
FUNCTION "SCALE_D" : Real   // FC334, SCL
TITLE = SCALE_D
{ S7_Optimized_Access := 'FALSE' }
AUTHOR : hugo
FAMILY : SIGPRO
NAME : SCALED
VERSION : 1.2
// Scale_D is used to translate and scale a DWORD input x to a real output.
// the input is limited to I_LO <= X <= I_HI.
   VAR_INPUT
      X : DWord;
      I_LO : DWord;
      I_HI : DWord;
      O_LO : Real;
      O_HI : Real;
   END_VAR
BEGIN


     IF #I_HI = #I_LO THEN
       #SCALE_D := #O_LO;
     ELSE
       #SCALE_D := (#O_HI - #O_LO) / DINT_TO_REAL(DWORD_TO_DINT(#I_HI) - DWORD_TO_DINT(#I_LO))
                  * DINT_TO_REAL(LIMIT(MN:=DWORD_TO_DINT(#I_LO),IN:=DWORD_TO_DINT(#X),MX:=DWORD_TO_DINT(#I_HI)) 
                  - DWORD_TO_DINT(#I_LO)) + #O_LO;
     END_IF;


   (* revision history
   hm  18. may. 2008 rev 1.0
     original version

   hm  13. nov. 2008 rev 1.1
     corrected formula for negative gradient

   hm  11. jan 2011  rev 1.2
     avoid division by 0
   *)
END_FUNCTION

FUNCTION "SCALE_R" : Real   // FC335, SCL
TITLE = SCALE_R
{ S7_Optimized_Access := 'FALSE' }
AUTHOR : hugo
FAMILY : SIGPRO
NAME : SCALER
VERSION : 1.2
// Scale_R is used to translate and scale a REAL input x to a real output.
// the input is limited to I_LO <= X <= I_HI.
   VAR_INPUT
      X : Real;
      I_LO : Real;
      I_HI : Real;
      O_LO : Real;
      O_HI : Real;
   END_VAR
BEGIN


     IF #I_LO = #I_HI THEN
       #SCALE_R := #O_LO;
     ELSE
       #SCALE_R := (#O_HI - #O_LO) / (#I_HI - #I_LO) * (LIMIT(MN:=#I_LO,IN:=#X,MX:=#I_HI) - #I_LO) + #O_LO;
     END_IF;


   (* revision history
   hm  18. may. 2008 rev 1.0
     original version

   hm  13. nov. 2008 rev 1.1
     corrected formula for negative gradient

   hm  11. jan 2011  rev 1.2
     avoid division by 0

   *)
END_FUNCTION

FUNCTION "SCALE_X2" : Real   // FC336, SCL
TITLE = SCALE_X2
{ S7_Optimized_Access := 'FALSE' }
AUTHOR : hugo
FAMILY : SIGPRO
NAME : SCALEX2
VERSION : 1.1
// this functiob block can scale up to two inputs.
// the input can select between two ues with true or false.
// the summed output is then scaled by an scale input K and a offset O can be added to the output.
// the min and max input configurations can be edited in the cfc editor by double clicking the symbol body.
   VAR_INPUT
      IN1 : Bool;
      IN2 : Bool;
      K : Real;
      O : Real;
      IN1_MIN : Real;
      IN1_MAX : Real;
      IN2_MIN : Real;
      IN2_MAX : Real;
   END_VAR
BEGIN


   #SCALE_X2 := (SEL(G:=#IN1,IN0:=#IN1_MIN, IN1:=#IN1_MAX)+ 
                SEL(G:=#IN2,IN0:=#IN2_MIN, IN1:=#IN2_MAX))*#K + #O;


   (* revision history
   hm  19. jan, 2007   rev 1.0
       original version

   hm  26. oct. 2008   rev 1.1
       code optimized

   *)
END_FUNCTION

FUNCTION "SCALE_X4" : Real   // FC337, SCL
TITLE = SCALE_X4
{ S7_Optimized_Access := 'FALSE' }
AUTHOR : hugo
FAMILY : SIGPRO
NAME : SCALEX4
VERSION : 1.0
// this function can scale up to 4 inputs.
// the input can select between two ues with true or false.
// the summed output is then scaled by an scale input K and a offset O can be added to the output.
// the min and max input configurations can be edited in the cfc editor by double clicking the symbol body.
   VAR_INPUT
      in1 : Bool;
      in2 : Bool;
      in3 : Bool;
      in4 : Bool;
      K : Real;
      O : Real;
      in1_min : Real;
      in1_max : Real;
      in2_min : Real;
      in2_max : Real;
      in3_min : Real;
      in3_max : Real;
      in4_min : Real;
      in4_max : Real;
   END_VAR
BEGIN


     IF NOT #in1 THEN #SCALE_X4 := #in1_min; ELSE #SCALE_X4 := #in1_max; END_IF;
     IF NOT #in2 THEN #SCALE_X4 := #SCALE_X4 + #in2_min; ELSE #SCALE_X4 := #SCALE_X4 + #in2_max; END_IF;
     IF NOT #in3 THEN #SCALE_X4 := #SCALE_X4 + #in3_min; ELSE #SCALE_X4 := #SCALE_X4 + #in3_max; END_IF;
     IF NOT #in4 THEN #SCALE_X4 := #SCALE_X4 + #in4_min; ELSE #SCALE_X4 := #SCALE_X4 + #in4_max; END_IF;
     #SCALE_X4 := #SCALE_X4 * #K + #O;

   (* revision history

   *)
END_FUNCTION

FUNCTION "SCALE_X8" : Real   // FC338, SCL
TITLE = SCALE_X8
{ S7_Optimized_Access := 'FALSE' }
AUTHOR : hugo
FAMILY : SIGPRO
NAME : SCALEX8
VERSION : 1.2
// this function can scale up to 4 inputs.
// the input can select between two ues with true or false.
// the summed output is then scaled by an scale input K and a offset O can be added to the output.
// the min and max input configurations can be edited in the cfc editor by double clicking the symbol body.
   VAR_INPUT
      in1 : Bool;
      in2 : Bool;
      in3 : Bool;
      in4 : Bool;
      in5 : Bool;
      in6 : Bool;
      in7 : Bool;
      in8 : Bool;
      K : Real;
      O : Real;
      in1_min : Real;
      in1_max : Real;
      in2_min : Real;
      in2_max : Real;
      in3_min : Real;
      in3_max : Real;
      in4_min : Real;
      in4_max : Real;
      in5_min : Real;
      in5_max : Real;
      in6_min : Real;
      in6_max : Real;
      in7_min : Real;
      in7_max : Real;
      in8_min : Real;
      in8_max : Real;
   END_VAR
BEGIN


   #SCALE_X8 := (SEL(G:=#in1,IN0:=#in1_min,IN1:=#in1_max) + 
                SEL(G:=#in2,IN0:=#in2_min,IN1:=#in2_max) + 
                SEL(G:=#in3,IN0:=#in3_min,IN1:=#in3_max) + 
                SEL(G:=#in4,IN0:=#in4_min,IN1:=#in4_max) +
                SEL(G:=#in5,IN0:=#in5_min,IN1:=#in5_max) + 
                SEL(G:=#in6,IN0:=#in6_min,IN1:=#in6_max) + 
                SEL(G:=#in7,IN0:=#in7_min,IN1:=#in7_max) + 
                SEL(G:=#in8,IN0:=#in8_min,IN1:=#in8_max))* #K + #O;


   (* revision history
   hm  19. jan. 2008   rev 1.0
       original version

   hm  26. oct. 2008   rev 1.1
       optimized code

   hm  24. jan. 2008   rev 1.2
       corrected error in formula
   *)
END_FUNCTION

FUNCTION "STAIR" : Real   // FC339, SCL
TITLE = STAIR
{ S7_Optimized_Access := 'FALSE' }
AUTHOR : oscat
FAMILY : SIGPRO
NAME : STAIR
VERSION : 1.4
// the function stair converts an anlog input signal to a staircase like output.
// D is the step width for the output signal.
// if D = 0 then the output follows the input without a chage.
   VAR_INPUT
      X : Real;
      D : Real;
   END_VAR
BEGIN


   IF #D > 0.0 THEN
       #STAIR := DINT_TO_REAL(REAL_TO_DINT(#X / #D)) * #D;
   ELSE
       #STAIR := #X;
   END_IF;


   (* revision history
   hm  28 jan 2007     rev 1.0
       original version

   hm  27 dec 2007     rev 1.1
       changed code for better performance

   hm  6. jan 2008     rev 1.2
       further performance improvement

   hm  26. oct. 2008       rev 1.3
       optimized code

   hm  10. mar. 2009   rev 1.4
       real constants updated to new systax using dot

   *)
END_FUNCTION

FUNCTION "WORD_TO_RANGE" : Real   // FC340, SCL
TITLE = WORD_TO_RANGE
{ S7_Optimized_Access := 'FALSE' }
AUTHOR : hugo
FAMILY : SIGPRO
NAME : WO2RA
VERSION : 1.1
// Word_to_Range converts a Byte into a real between low and high.
   VAR_INPUT
      X : Word;
      low : Real;
      high : Real;
   END_VAR
BEGIN


   #WORD_TO_RANGE := (#high - #low) * DINT_TO_REAL(WORD_TO_DINT(#X)) * 0.00001525902189669640 + #low;


   (* revision history
   hm  9. jan 2008 rev 1.0
       original version

   hm  10. mar. 2009   rev 1.1
       improved code
   *)
END_FUNCTION

// ===== PLC "Engineering automation"  Unspecific CPU S7 300 =====

VAR_GLOBAL CONSTANT   // PLC tag table "STEP7 classic symbols"
   "debug" : Bool := FALSE;
   "N" : Int := 0;
   "offset" : Int := 0;
   "one" : Byte := 16#01;
   "offset_1" : DWord := 0;
END_VAR

DATA_BLOCK "IDB_STIME"   // DB64
{ S7_Optimized_Access := 'FALSE' }
AUTHOR : dalbi
FAMILY : MEASURE
VERSION : 0.0
// stored: InstanceOfName STIME
"STIME"
BEGIN
END_DATA_BLOCK

FUNCTION_BLOCK "STIME"   // FB64, SCL
TITLE = STIME
{ S7_Optimized_Access := 'FALSE' }
AUTHOR : dalbi
FAMILY : MEASURE
NAME : STIME
VERSION : 1.4
// this function block makes sure that the timer of a siemens sps counts from 0 - 2^32-1.
   VAR_OUTPUT
      tx : DWord;
      at_tx AT tx : Array[0..31] of Bool;
   END_VAR
   VAR
      last_time : DWord;
      bit31 : Bool;
      init : Bool := TRUE;
   END_VAR
   VAR_TEMP
      TOP_SI : Struct
         EV_CLASS : Byte;
         EV_NUM : Byte;
         PRIORITY : Byte;
         NUM : Byte;
         TYP2_3 : Byte;
         TYP1 : Byte;
         ZI1 : Word;
         ZI2_3 : DWord;
      END_STRUCT;
      START_UP_SI : Struct
         EV_CLASS : Byte;
         EV_NUM : Byte;
         PRIORITY : Byte;
         NUM : Byte;
         TYP2_3 : Byte;
         TYP1 : Byte;
         ZI1 : Word;
         ZI2_3 : DWord;
      END_STRUCT;
      ERR : Int;
   END_VAR
BEGIN


   (* this FB is only necessary for siemens sps
   the siemens sps timer counts from 0 to 2^31-1 and starts at 0 sfter overrun.
   this means that the bit 31 (the highest bit ) will never be used and therefore
   a problem arises when t2 - t1 is checked.
   t2 - t1 is always valid also in an timer overrun situation where the time t1 is very high and t2 is very low.
   the result of the subtraction t2 - t1 however is still valid.
   this calculation does not work for soiemens because the highest bit is not used.

   this module stores the highest bit, changes the highest bit at every overrun occurence and stuffs ther highest bit in the output.
   the output is then used by t_plc_us and t_plc_ms.

   the correction needs and fb and not a function because the value of the highest bit has to be stored.

   do never use this function block in a codesys environment. the timer in codesys is correct and runs from 0 to 2^32-1
   *)

   (* read actual startup info *)
   (* OB1_SCAN_1  BYTE  -  B#16#01: Abschluss des Neustarts (Warmstarts)
                        -  B#16#02: Abschluss des Wiederanlaufs
                        -  B#16#03: Abschluss des freien Zyklus
                        -  B#16#04: Abschluss des Kaltstarts
                        -  B#16#05: Erster OB 1-Zyklus der neuen Master-CPU nach 
                                    Master-Reserve-Umschaltung und STOP des 
                                    bisherigen Masters *)

   #ERR := RD_SINFO (TOP_SI => #TOP_SI, START_UP_SI => #START_UP_SI);

   (* reset last_time on system startup *)
   IF #TOP_SI.EV_NUM = 1 OR #TOP_SI.EV_NUM = 2 OR #TOP_SI.EV_NUM = 4 OR NOT #init THEN 
       #last_time := 0;
       #bit31 := false;
       #init := true;
   END_IF;

   (* read the system timer *)
   #tx := DINT_TO_DWORD(T_CONV(TIME_TCK()));

   (* check for overrun *)
   IF DWORD_TO_DINT(#tx) < DWORD_TO_DINT(#last_time) THEN
       (* an overrun has occured, change the value of the highest bit *)
       #bit31 := NOT #bit31;
   END_IF;

   (* stuff the highest bit into the timer value *)
   #at_tx[7] := #bit31;

   (* remember the last system time for the next overrun check *)
   #last_time := #tx;


   (* revision history
   DA  14.9.2007 rev 1.0
     original version

   DA  24.2.2008 rev 1.1
     added self reset on system startup

   DA   2.5.2008 rev 1.2
     corect a problem running under OB35

   DA  12.3.2009 rev 1.3
     corect a problem run on different CPUs

   DA  22.12.2009 rev 1.4
     corect a problem on startup
   *)
END_FUNCTION_BLOCK

FUNCTION_BLOCK "TP_1D"   // FB68, SCL
TITLE = TP_1D
{ S7_Optimized_Access := 'FALSE' }
AUTHOR : hugo
FAMILY : GENERAT
NAME : TP_1D
VERSION : 1.0
// TP_2 generates a pulse every time it is calles with in := TRUE.
// the module will reset IN by itself so no clearing of in is necessary.
// in addition the timer can be cleared asynchronously with rst.
// also the rst input is cleared by the module itself.
// the timer can be retriggered as often as necessary. it will count PT from the last trigger.
// after the time PT1 is elapsed, the timer blocks itself for PT2 and only allow new sequences after PT2 has elapsed.
// 
// uses: T_PLC_MS [FC64]
//       STIME [FB64],IDB_STIME [DB64]
   VAR_INPUT
      IN : Bool;
      PT1 : Time;
      PTD : Time;
      RST : Bool;
   END_VAR
   VAR_OUTPUT
      Q : Bool;
      W : Bool;
   END_VAR
   VAR
      tx : Time;
      start : Time;
      ix : Bool;
   END_VAR
BEGIN


   (* read system timer *)
   #tx := T_CONV(DWORD_TO_DINT("T_PLC_MS"()));

   IF #RST THEN
       #Q := FALSE;
       #RST := FALSE;
       #W := FALSE;
   ELSIF #W THEN
       IF #tx - #start >= #PTD THEN
           #W := FALSE;
       END_IF;
   ELSIF #IN AND NOT #ix THEN
       #Q := TRUE;
       #start := #tx;
       #IN := FALSE;
   ELSIF #tx - #start >= #PT1 THEN
       #Q := FALSE;
       #W := TRUE;
       #start := #tx;
   END_IF;

   #ix := #IN;



   (* revision history
   hm  28. jun. 2008
       original version

   *)
END_FUNCTION_BLOCK

FUNCTION_BLOCK "TC_S"   // FB134, SCL
TITLE = TC_S
{ S7_Optimized_Access := 'FALSE' }
AUTHOR : hugo
FAMILY : MEASURE
NAME : TC_S
VERSION : 1.2
// TC_S delivers the time it was last called on the output TC in seconds.
// 
// uses: T_PLC_US [FC65]
//       STIME [FB64],IDB_STIME [DB64]
   VAR_OUTPUT
      TC : Real;
   END_VAR
   VAR
      init : Bool;
      tx : DWord;
      last : DWord;
   END_VAR
   VAR_TEMP
      TOP_SI : Struct
         EV_CLASS : Byte;
         EV_NUM : Byte;
         PRIORITY : Byte;
         NUM : Byte;
         TYP2_3 : Byte;
         TYP1 : Byte;
         ZI1 : Word;
         ZI2_3 : DWord;
      END_STRUCT;
      START_UP_SI : Struct
         EV_CLASS : Byte;
         EV_NUM : Byte;
         PRIORITY : Byte;
         NUM : Byte;
         TYP2_3 : Byte;
         TYP1 : Byte;
         ZI1 : Word;
         ZI2_3 : DWord;
      END_STRUCT;
      ERR : Int;
   END_VAR
BEGIN


   (* read actual startup info *)
   (* OB1_SCAN_1  BYTE  -  B#16#01: Abschluss des Neustarts (Warmstarts)
                        -  B#16#02: Abschluss des Wiederanlaufs
                        -  B#16#03: Abschluss des freien Zyklus
                        -  B#16#04: Abschluss des Kaltstarts
                        -  B#16#05: Erster OB 1-Zyklus der neuen Master-CPU nach 
                                    Master-Reserve-Umschaltung und STOP des 
                                    bisherigen Masters *)

     #ERR := RD_SINFO (TOP_SI => #TOP_SI, START_UP_SI => #START_UP_SI);

   (* reset last_time on system startup *)
   IF #TOP_SI.EV_NUM = 1 OR #TOP_SI.EV_NUM = 2 OR #TOP_SI.EV_NUM = 4 THEN 
       #last := 0;
       #init := FALSE;
   END_IF;

   (* read system timer *)
   #tx := "T_PLC_US"();

   IF NOT #init THEN
       #init := TRUE;
       #TC := 0.0;
   ELSE
       #TC := (DINT_TO_REAL(DWORD_TO_DINT(#tx)) - DINT_TO_REAL(DWORD_TO_DINT(#last)))*1.0E-6;
   END_IF;
   #last := #tx;


   (* revision history
   hm  13. mar. 2008   rev 1.0
       original version

   hm  16. mar 2008    rev 1.1
       added type conversion to avoid warnings under codesys 3.0

   hm  11. mar. 2009   rev 1.2
       changed real constants to use dot syntax

   *)
END_FUNCTION_BLOCK

FUNCTION_BLOCK "DRIVER_1"   // FB202, SCL
TITLE = DRIVER_1
{ S7_Optimized_Access := 'FALSE' }
AUTHOR : hugo
FAMILY : AUTOMAT
NAME : DRIVER_1
VERSION : 1.0
// driver_1 is a multi purpose driver.
// a rising edge in in sets the output high if toggle is flase. while toggle is true, a rising edge on in toggles the output Q.
// if a timeout is specified the output q will be reset to false automatically after the timeout has elapsed.
// a asynchronous reset and set will force the output high or low respectively.
   VAR_INPUT
      Toggle_Mode : Bool;
      Timeout : Time;
      SET : Bool;
      IN : Bool;
      RST : Bool;
   END_VAR
   VAR_OUTPUT
      Q : Bool;
   END_VAR
   VAR
      off : TON;
      edge : Bool;
   END_VAR
BEGIN


     IF #off.Q THEN #Q := FALSE; END_IF;
     IF #RST THEN
       #Q := FALSE;
     ELSIF #SET THEN
       #Q := TRUE;
     ELSIF #IN AND NOT #edge THEN
       IF #Toggle_Mode THEN #Q := NOT #Q; ELSE #Q := TRUE; END_IF;
     END_IF;
     #edge := #IN;
     IF #Timeout > t#0s THEN #off(IN := #Q, PT := #Timeout); END_IF;


   (* revision history
   hm  2. jan 2008   rev 1.0
     original version

   *)
END_FUNCTION_BLOCK

FUNCTION_BLOCK "DRIVER_4"   // FB203, SCL
TITLE = DRIVER_4
{ S7_Optimized_Access := 'FALSE' }
AUTHOR : hugo
FAMILY : AUTOMAT
NAME : DRIVER_4
VERSION : 1.0
// driver_1 is a multi purpose driver.
// a rising edge in in sets the output high if toggle is flase. while toggle is true, a rising edge on in toggles the output Q.
// if a timeout is specified the output q will be reset to false automatically after the timeout has elapsed.
// a asynchronous reset and set will force the output high or low respectively.
// 
// uses: DRIVER_1 [FB202]
   VAR_INPUT
      Toggle_Mode : Bool;
      Timeout : Time;
      SET : Bool;
      IN0 : Bool;
      IN1 : Bool;
      IN2 : Bool;
      IN3 : Bool;
      RST : Bool;
   END_VAR
   VAR_OUTPUT
      Q0 : Bool;
      Q1 : Bool;
      Q2 : Bool;
      Q3 : Bool;
   END_VAR
   VAR
      d0 : "DRIVER_1";
      d1 : "DRIVER_1";
      d2 : "DRIVER_1";
      d3 : "DRIVER_1";
   END_VAR
BEGIN


     #d0(SET:=#SET, IN:=#IN0, RST:=#RST, Toggle_Mode:=#Toggle_Mode, Timeout:=#Timeout);
     #d1(SET:=#SET, IN:=#IN1, RST:=#RST, Toggle_Mode:=#Toggle_Mode, Timeout:=#Timeout);
     #d2(SET:=#SET, IN:=#IN2, RST:=#RST, Toggle_Mode:=#Toggle_Mode, Timeout:=#Timeout);
     #d3(SET:=#SET, IN:=#IN3, RST:=#RST, Toggle_Mode:=#Toggle_Mode, Timeout:=#Timeout);
     #Q0 := #d0.Q;
     #Q1 := #d1.Q;
     #Q2 := #d2.Q;
     #Q3 := #d3.Q;


   (* revision history
   hm  2. jan 2008   rev 1.0
     original version

   *)
END_FUNCTION_BLOCK

FUNCTION_BLOCK "FLOW_CONTROL"   // FB204, SCL
TITLE = FLOW_CONTROL
{ S7_Optimized_Access := 'FALSE' }
AUTHOR : hugo
FAMILY : AUTOMAT
NAME : FLOWCTR
VERSION : 1.0
// FLOW_CONTROL switches a valves depending on the input in.
// flow control also limits the maximum ontime of the valve and controls pressure on the output side.
// 
// uses: TP_1D [FB68]
//       T_PLC_MS [FC64] 
//       STIME [FB64],IDB_STIME [DB64]
   VAR_INPUT
      IN : Bool;
      REQ : Bool;
      ENQ : Bool;
      RST : Bool;
      T_AUTO : Time := T#1H;
      T_DELAY : Time := T#23H;
   END_VAR
   VAR_OUTPUT
      Q : Bool;
      STATUS : Byte;
   END_VAR
   VAR
      _timer : "TP_1D";
   END_VAR
BEGIN


   #STATUS := 100;
   IF #RST THEN
       #Q := FALSE;
       #_timer(RST := TRUE);
       #_timer.RST := FALSE;
       #STATUS := 103;
   ELSIF #ENQ THEN
       IF #IN THEN
           #STATUS := 101;
       END_IF;
       IF #REQ THEN
           (* timer will generate a timed pulse after TP goes high *)
           #_timer.PT1 := #T_AUTO;
           #_timer.PTD := #T_DELAY;
           #_timer.IN := TRUE;
           #STATUS := 102;
       END_IF;
   END_IF;


   (* set output and run timer *)
   #_timer();
   #_timer.IN := FALSE;
   #Q := (#IN AND #ENQ) OR #_timer.Q;



   (* revision history
   hm  28. jun. 2008   rev 1.0
       original version

   *)
END_FUNCTION_BLOCK

FUNCTION_BLOCK "FT_PROFILE"   // FB206, SCL
TITLE = FT_PROFILE
{ S7_Optimized_Access := 'FALSE' }
AUTHOR : tobias
FAMILY : AUTOMAT
NAME : FT_PROF
VERSION : 1.1
// FT_Profile generates an output signal which is defined by values over a time scale.
// the different values are connected by ramps between the individual values.
// a rising edge on E starts the output signal generation and E = True can delay time_3 / value_3 as long as it stays true.
// an additional multiplier K can be used to multiply the output and an offset O can be added to the output dynamically.
// 
// uses: T_PLC_MS [FC64]
//       STIME [FB64],IDB_STIME [DB64]
//       MULTIME [FC203]
   VAR_INPUT
      K : Real := 1.0e+0;
      O : Real;
      "M" : Real := 1.0e+0;
      "E" : Bool;
      value_0 : Real;
      time_1 : Time;
      value_1 : Real;
      time_2 : Time;
      value_2 : Real;
      time_3 : Time;
      value_3 : Real;
      time_10 : Time;
      value_10 : Real;
      time_11 : Time;
      value_11 : Real;
      time_12 : Time;
      value_12 : Real;
      time_13 : Time;
      value_13 : Real;
   END_VAR
   VAR_OUTPUT
      Y : Real;
      RUN : Bool;
      ET : Time;
   END_VAR
   VAR
      tx : Time;
      edge : Bool;
      state : Byte;
      ta : Time;
      tb : Time;
      t_0 : Time;
      temp : Real;
      va : Real;
      vb : Real;
   END_VAR
BEGIN


     (* read system time *)
     #tx := T_CONV(DWORD_TO_DINT("T_PLC_MS"()));

     (* determine start condition *)
     IF #"E" AND NOT #edge THEN
         #RUN := TRUE;
         #ET := t#0s;
         #t_0 := #tx;
         #ta := #tx;
         #tb := "MULTIME"(t:=#time_1,M:=#"M");
         #va := #value_0;
         #vb := #value_1;
         #temp := #value_0;
         #state := 1;
     END_IF;
     #edge := #"E";

     (* generate startup profile *)
     IF #RUN THEN
         CASE BYTE_TO_INT(#state) OF
             1:    IF #tx - #ta >= #tb THEN
                     #ta := #ta + #tb;
                     #tb := "MULTIME"(t:=#time_2 - #time_1,M:=#"M");
                     #va := #value_1;
                     #vb := #value_2;
                     #temp := #value_1;
                     #state := 2;
                 ELSE
                     #temp := ((#vb - #va) * DINT_TO_REAL(T_CONV(#tx - #ta)) / DINT_TO_REAL(T_CONV(#tb)) + #va);
                 END_IF;
             2:    IF #tx - #ta >= #tb THEN
                     #ta := #ta + #tb;
                     #tb := "MULTIME"(t:=#time_3 - #time_2,M:=#"M");
                     #va := #value_2;
                     #vb := #value_3;
                     #temp := #value_2;
                     #state := 3;
                 ELSE
                     #temp := ((#vb - #va) * DINT_TO_REAL(T_CONV(#tx - #ta)) / DINT_TO_REAL(T_CONV(#tb)) + #va);
                 END_IF;
             3:    IF #tx - #ta >= #tb THEN
                     #ta := #ta + #tb;
                     #tb := "MULTIME"(t:=#time_10 - #time_3,M:=#"M");
                     #va := #value_3;
                     #vb := #value_10;
                     #temp := #value_3;
                     #state := 4;
                 ELSE
                     #temp := ((#vb - #va) * DINT_TO_REAL(T_CONV(#tx - #ta)) / DINT_TO_REAL(T_CONV(#tb)) + #va);
                 END_IF;
             4 :    IF #tx - #ta >= #tb THEN
                     #ta := #ta + #tb;
                     #tb := "MULTIME"(t:=#time_11 - #time_10,M:=#"M");
                     #va := #value_10;
                     #vb := #value_11;
                     #temp := #value_10;
                     IF #"E" THEN #state := 5; ELSE #state := 6; END_IF;
                 ELSE
                     #temp := ((#vb - #va) * DINT_TO_REAL(T_CONV(#tx - #ta)) / DINT_TO_REAL(T_CONV(#tb)) + #va);
                 END_IF;
             5:    (* extend the signal while E is true *)
                 IF #"E" THEN
                     #ta := #tx;
                 ELSE
                     #state := 6;
                 END_IF;
             6:    IF #tx - #ta >= #tb THEN
                     #ta := #ta + #tb;
                     #tb := "MULTIME"(t:=#time_12 - #time_11,M:=#"M");
                     #va := #value_11;
                     #vb := #value_12;
                     #temp := #value_11;
                     #state := 7;
                 ELSE
                     #temp := ((#vb - #va) * DINT_TO_REAL(T_CONV(#tx - #ta)) / DINT_TO_REAL(T_CONV(#tb)) + #va);
                 END_IF;
             7:    IF #tx - #ta >= #tb THEN
                     #ta := #ta + #tb;
                     #tb := "MULTIME"(t:=#time_13 - #time_12,M:=#"M");
                     #va := #value_12;
                     #vb := #value_13;
                     #temp := #value_12;
                     #state := 8;
                 ELSE
                     #temp := ((#vb - #va) * DINT_TO_REAL(T_CONV(#tx - #ta)) / DINT_TO_REAL(T_CONV(#tb)) + #va);
                 END_IF;
             8:    IF #tx - #ta >= #tb THEN
                     #temp := #value_13;
                     #RUN := FALSE;
                 ELSE
                     #temp := ((#vb - #va) * DINT_TO_REAL(T_CONV(#tx - #ta)) / DINT_TO_REAL(T_CONV(#tb)) + #va);
                 END_IF;
         END_CASE;
         #Y := #temp * #K + #O;
         #ET := #tx - #t_0;
     END_IF;

   (* revision history
   hm  27 feb 2007    rev 1.0
     original version

   hm  15. sep2007    rev 1.1
     replaced Time() with T_PLC_MS for compatibility and performance reasons

   *)
END_FUNCTION_BLOCK

FUNCTION_BLOCK "INC_DEC"   // FB207, SCL
TITLE = INC_DEC
{ S7_Optimized_Access := 'FALSE' }
AUTHOR : oscat
FAMILY : AUTOMAT
NAME : INC_DEC
VERSION : 1.0
// incremental decoder with quadruple accuracy.
// 2 pulses for each channel are created for each directional pulse.
   VAR_INPUT
      CHa : Bool;
      CHb : Bool;
      RST : Bool;
   END_VAR
   VAR_OUTPUT
      dir : Bool;
      cnt : Int;
   END_VAR
   VAR
      edgea : Bool;
      clk : Bool;
      clka : Bool;
      clkb : Bool;
      edgeb : Bool;
      axb : Bool;
   END_VAR
BEGIN


     #axb := #CHa XOR #CHb;

     (* create pulses for channel a *)
     #clka := #CHa XOR #edgea;
     #edgea := #CHa;

     #clkb := #CHb XOR #edgeb;
     #edgeb := #CHb;

     (* create pulses for both channels *)
     #clk := #clka OR #clkb;

     (* set the direction output *)
     IF #axb AND #clka THEN #dir := TRUE; END_IF;
     IF #axb AND #clkb THEN #dir := FALSE; END_IF;

     (* increment or decrement the counter *)
     IF #clk AND #dir THEN #cnt := #cnt + 1; END_IF;
     IF #clk AND NOT #dir THEN #cnt := #cnt -1; END_IF;

     (* reset the counter if rst active *)
     IF #RST THEN #cnt := 0; END_IF;
END_FUNCTION_BLOCK

FUNCTION_BLOCK "INTERLOCK"   // FB208, SCL
TITLE = INTERLOCK
{ S7_Optimized_Access := 'FALSE' }
AUTHOR : hugo
FAMILY : AUTOMAT
NAME : INTLOCK
VERSION : 1.0
// INTERLOCK has two inputs I1 and I2 which drive the corresponding outputs Q1 and Q2.
// the inputs signals lock each other out and therfore I1 can only drive Q1 when I2 is Low and vice versa.
// The input TL specifies a dead time between two outputs can become active.
// an output can only become active when the other output was not active for the time TL.
   VAR_INPUT
      I1 : Bool;
      I2 : Bool;
      TL : Time;
   END_VAR
   VAR_OUTPUT
      Q1 : Bool;
      Q2 : Bool;
   END_VAR
   VAR
      T_1 : TOF;
      T_2 : TOF;
   END_VAR
BEGIN


     (* the input signal have a run delay to lockout the other input *)
     #T_1(IN := #I1, PT := #TL);
     #T_2(IN := #I2, PT := #TL);

     #Q1 := #I1 AND NOT #T_2.Q;
     #Q2 := #I2 AND NOT #T_1.Q;


   (* revision history

   hm  28 sep 2007    rev 1.0
     original version

   *)
END_FUNCTION_BLOCK

FUNCTION_BLOCK "INTERLOCK_4"   // FB209, SCL
TITLE = INTERLOCK_4
{ S7_Optimized_Access := 'FALSE' }
AUTHOR : hugo
FAMILY : AUTOMAT
NAME : INTLOCK4
VERSION : 1.1
// INTERLOCK_4 detects one of 4 switches and delivers the number of the switch pressed on the output out
// a output tp is true for one cycle if the output has changed.
// a setup variable MODE selects between 3 different modes:
// MODE = 0, any input active will disable all other inputs
// MODE = 1, the input with the highest number will be acepted
// mode = 2, the input last pressed will disable all others
   VAR_INPUT
      I0 : Bool;
      I1 : Bool;
      I2 : Bool;
      I3 : Bool;
      "E" : Bool;
      MODE : Int;
   END_VAR
   VAR_OUTPUT
      OUT : Byte;
      TP : Bool;
   END_VAR
   VAR
      in : Byte;
      _in AT in : Array[0..7] of Bool;
      last : Byte;
      _last AT last : Array[0..7] of Bool;
      old : Byte;
      lmode : Int;
   END_VAR
BEGIN


   (* check if enable is active *)
   IF #"E" THEN
   (* reset all vars when there is a mode change on thy fly *)
       IF #MODE <> #lmode THEN
           #OUT := 0;
           #last := 0;
           #old := 0;
           #lmode := #MODE;
       END_IF;
       (* load inputs into in *)
       #_in[0] := #I0; 
       #_in[1] := #I1; 
       #_in[2] := #I2; 
       #_in[3] := #I3;
       (* only execute when there is any change *)
       IF #in <> #last THEN
           (* only execute when inputs have chages state *)
           CASE #MODE OF
               0:  (* output directly display inputs as bits in byte out *)
                   #OUT := #in;

               1:  (* the input with the highest number will be acepted *)
                   IF #_in[3] THEN #OUT := 8;
                   ELSIF #_in[2] THEN #OUT := 4;
                   ELSIF #_in[1] THEN #OUT := 2;
                   ELSE #OUT := #in;
                   END_IF;

               2:  (* input last pressed will be displayed only *)
                   #last := ((#in XOR #last) AND #in);
                   IF #_last[3] THEN #OUT := 8;
                   ELSIF #_last[2] THEN #OUT := 4;
                   ELSIF #_last[1] THEN #OUT := 2;
                   ELSE #OUT := #last;
                   END_IF;

               3:  (* any input active will disable all other inputs *)
                   IF (#OUT AND #in) = 0 THEN
                       IF #_in[3] THEN #OUT := 8;
                       ELSIF #_in[2] THEN #OUT := 4;
                       ELSIF #_in[1] THEN #OUT := 2;
                       ELSE #OUT := #in;
                       END_IF;
                   END_IF;

           END_CASE;
           #last := #in;
       END_IF;
       #TP := #OUT <> #old;
       #old := #OUT;
   ELSE
       #OUT := 0;
       #last := 0;
       #old := 0;
       #lmode := 0;
       #TP := FALSE;
   END_IF;


   (* revision history
   hm  24. oct 2008    rev 1.0
       original version

   hm  14. mar. 2009   rev 1.1
       replaced double assignments

   *)
END_FUNCTION_BLOCK

FUNCTION_BLOCK "MANUAL_1"   // FB210, SCL
TITLE = MANUAL_1
{ S7_Optimized_Access := 'FALSE' }
AUTHOR : hugo
FAMILY : AUTOMAT
NAME : MANUAL1
VERSION : 1.2
// MANUAL_1 is a manual override for digital signals.
// When MAN = FALSE, the output follows IN and when MAN = TRUE the Output follows M_I.
   VAR_INPUT
      IN : Bool;
      MAN : Bool;
      M_I : Bool;
      SET : Bool;
      RST : Bool;
   END_VAR
   VAR_OUTPUT
      Q : Bool;
      STATUS : Byte;
   END_VAR
   VAR
      S_edge : Bool;
      r_edge : Bool;
      edge : Bool;
   END_VAR
BEGIN


   IF NOT #MAN THEN
       #Q := #IN;
       #STATUS := 100;
       #edge := FALSE;
   ELSIF NOT #S_edge AND #SET THEN
       #Q := TRUE;
       #edge := TRUE;
       #STATUS := 101;
   ELSIF NOT #r_edge AND #RST THEN
       #Q := FALSE;
       #edge := TRUE;
       #STATUS := 102;
   ELSIF NOT #edge THEN
       #Q := #M_I;
       #STATUS := 103;
   END_IF;

   (* remember levels of manual signals *)
   #S_edge := #SET;
   #r_edge := #RST;


   (* revision history
   hm  17. jun 2008    rev 1.0
       original version

   hm  17. oct 2008    rev 1.1
       deleted unnecessary variable m_edge

   hm  14. mar. 2009   rev 1.2
       replaced double assignments

   *)
END_FUNCTION_BLOCK

FUNCTION_BLOCK "MANUAL_2"   // FB211, SCL
TITLE = MANUAL_2
{ S7_Optimized_Access := 'FALSE' }
AUTHOR : hugo
FAMILY : AUTOMAT
NAME : MANUAL2
VERSION : 1.0
// MANUAL_2 is a manual override for boolean signals.
// it has static force high and low as well as a manual input.
   VAR_INPUT
      IN : Bool;
      ENA : Bool;
      ON : Bool;
      OFF : Bool;
      MAN : Bool;
   END_VAR
   VAR_OUTPUT
      Q : Bool;
      STATUS : Byte;
   END_VAR
BEGIN


   IF #ENA THEN
       IF NOT #ON AND NOT #OFF THEN
           #Q := #IN;
           #STATUS := 100;
       ELSIF #ON AND NOT #OFF THEN
           #Q := TRUE;
           #STATUS := 101;
       ELSIF NOT #ON AND #OFF THEN
           #Q := FALSE;
           #STATUS := 102;
       ELSE
           #Q := #MAN;
           #STATUS := 103;
       END_IF;
   ELSE
       #Q := FALSE;
       #STATUS := 104;
   END_IF;



   (* revision history
   hm  22. sep. 2008       rev 1.0
       original version

   *)
END_FUNCTION_BLOCK

FUNCTION_BLOCK "MANUAL_4"   // FB212, SCL
TITLE = MANUAL_4
{ S7_Optimized_Access := 'FALSE' }
AUTHOR : hugo
FAMILY : AUTOMAT
NAME : MANUAL4
VERSION : 1.0
// MANUAL_4 is a manual override for digital signals.
// When MAN = FALSE, the output follows IN and when MAN = TRUE the Output follows M_I.
// 
// uses: INC [FC90]
   VAR_INPUT
      I0 : Bool;
      I1 : Bool;
      I2 : Bool;
      I3 : Bool;
      MAN : Bool;
      STP : Bool;
      M0 : Bool;
      M1 : Bool;
      M2 : Bool;
      M3 : Bool;
   END_VAR
   VAR_OUTPUT
      Q0 : Bool;
      Q1 : Bool;
      Q2 : Bool;
      Q3 : Bool;
      STATUS : Byte;
   END_VAR
   VAR
      edge : Bool;
      pos : Int;
      tog : Bool;
   END_VAR
BEGIN


   IF #MAN THEN
       IF NOT #tog THEN
           #Q0 := #M0;
           #Q1 := #M1;
           #Q2 := #M2;
           #Q3 := #M3;
           #STATUS := 101;
       END_IF;
       IF #STP AND NOT #edge THEN
           #tog := TRUE;
           CASE #pos OF
               0:  #Q0 := TRUE;
                   #Q1 := FALSE;
                   #Q2 := FALSE;
                   #Q3 := FALSE;
                   #STATUS := 110;
               1:  #Q0 := FALSE;
                   #Q1 := TRUE;
                   #Q2 := FALSE;
                   #Q3 := FALSE;
                   #STATUS := 111;
               2:  #Q0 := FALSE;
                   #Q1 := FALSE;
                   #Q2 := TRUE;
                   #Q3 := FALSE;
                   #STATUS := 112;
               3:  #Q0 := FALSE;
                   #Q1 := FALSE;
                   #Q2 := FALSE;
                   #Q3 := TRUE;
                   #STATUS := 113;
           END_CASE;
           #pos := "INC"(X:=#pos,D:=1,M:=3);
       END_IF;
   ELSE
       #Q0 := #I0;
       #Q1 := #I1;
       #Q2 := #I2;
       #Q3 := #I3;
       #STATUS := 100;
       #tog := FALSE;
       #pos := 0;
   END_IF;

   (* remember status of stp *)
   #edge := #STP;



   (* revision history
   hm  17. jun 2008        rev 1.0
       original version

   *)
END_FUNCTION_BLOCK

FUNCTION_BLOCK "PARSET"   // FB213, SCL
TITLE = PARSET
{ S7_Optimized_Access := 'FALSE' }
AUTHOR : hugo
FAMILY : AUTOMAT
NAME : PARSET
VERSION : 1.1
// parset selects on of 4 parameter sets adressed by the inputs A0 and A1. if TC is specified, the change of the outputs
// is ramped by the time tc
// 
// uses: T_PLC_MS [FC64]
//       STIME [FB64],IDB_STIME [DB64]
   VAR_INPUT
      A0 : Bool;
      A1 : Bool;
      X01 : Real;
      X02 : Real;
      X03 : Real;
      X04 : Real;
      X11 : Real;
      X12 : Real;
      X13 : Real;
      X14 : Real;
      X21 : Real;
      X22 : Real;
      X23 : Real;
      X24 : Real;
      X31 : Real;
      X32 : Real;
      X33 : Real;
      X34 : Real;
      TC : Time;
   END_VAR
   VAR_OUTPUT
      P1 : Real;
      P2 : Real;
      P3 : Real;
      P4 : Real;
   END_VAR
   VAR
      X : Array[0..3, 1..4] of Real;
      S1 : Real;
      S2 : Real;
      S3 : Real;
      S4 : Real;
      tx : DWord;
      last : DWord;
      start : Bool;
      set : Byte;
      _set AT set : Array[0..7] of Bool;
      init : Bool;
   END_VAR
BEGIN


     (* read system_time *)
     #tx := "T_PLC_MS"();

     (* init sequence *)
     IF NOT #init THEN
       #_set[0] := NOT #A0;
       #init := TRUE;
       #X[0,1] := #X01;
       #X[0,2] := #X02;
       #X[0,3] := #X03;
       #X[0,4] := #X04;
       #X[1,1] := #X11;
       #X[1,2] := #X12;
       #X[1,3] := #X13;
       #X[1,4] := #X14;
       #X[2,1] := #X21;
       #X[2,2] := #X22;
       #X[2,3] := #X23;
       #X[2,4] := #X24;
       #X[3,1] := #X31;
       #X[3,2] := #X32;
       #X[3,3] := #X33;
       #X[3,4] := #X34;
       #P1 := #X01;
       #P2 := #X02;
       #P3 := #X03;
       #P4 := #X04;
     END_IF;

     (* check for input change *)
     IF (#A0 XOR #_set[0]) OR (#A1 XOR #_set[1]) THEN
       (* a new set is selected *)
       #_set[0] := #A0;
       #_set[1] := #A1;
       IF #TC > t#0s THEN
         #start := TRUE;
         #last := #tx;
         (* save the step speed for the output changes in S *)
         #S1 := (#X[BYTE_TO_INT(#set),1] - #P1)/DINT_TO_REAL(T_CONV(#TC));
         #S2 := (#X[BYTE_TO_INT(#set),2] - #P2)/DINT_TO_REAL(T_CONV(#TC));
         #S3 := (#X[BYTE_TO_INT(#set),3] - #P3)/DINT_TO_REAL(T_CONV(#TC));
         #S4 := (#X[BYTE_TO_INT(#set),4] - #P4)/DINT_TO_REAL(T_CONV(#TC));
       END_IF;
     ELSIF #start AND DWORD_TO_DINT(#tx) - DWORD_TO_DINT(#last) < T_CONV(#TC) THEN
       (* ramp the outputs to the new value *)
       #P1 := #X[BYTE_TO_INT(#set),1] - #S1*(DINT_TO_REAL((T_CONV(#TC) - DWORD_TO_DINT(#tx) + DWORD_TO_DINT(#last))));
       #P2 := #X[BYTE_TO_INT(#set),2] - #S2*(DINT_TO_REAL((T_CONV(#TC) - DWORD_TO_DINT(#tx) + DWORD_TO_DINT(#last))));
       #P3 := #X[BYTE_TO_INT(#set),3] - #S3*(DINT_TO_REAL((T_CONV(#TC) - DWORD_TO_DINT(#tx) + DWORD_TO_DINT(#last))));
       #P4 := #X[BYTE_TO_INT(#set),4] - #S4*(DINT_TO_REAL((T_CONV(#TC) - DWORD_TO_DINT(#tx) + DWORD_TO_DINT(#last))));
     ELSE
       (* make sure outputs match the correct set values *)
       #start := FALSE;
       #P1 := #X[BYTE_TO_INT(#set),1];
       #P2 := #X[BYTE_TO_INT(#set),2];
       #P3 := #X[BYTE_TO_INT(#set),3];
       #P4 := #X[BYTE_TO_INT(#set),4];
     END_IF;

   (* revision history
   hm  2.11.2007       rev 1.0
       original version

   hm  16. mar. 2008   rev 1.1
       added type conversions to avoid warnings under codesys 3.0

   *)
END_FUNCTION_BLOCK

FUNCTION_BLOCK "PARSET2"   // FB214, SCL
TITLE = PARSET2
{ S7_Optimized_Access := 'FALSE' }
AUTHOR : hugo
FAMILY : AUTOMAT
NAME : PARSET2
VERSION : 1.0
// parset2 selects on of 4 parameter sets depending on the value of X. if TC is specified, the change of the outputs
// is ramped by the time TC
// 
// uses: PARSET [FB213]
//       T_PLC_MS [FC64] 
//       STIME [FB64],IDB_STIME [DB64]
   VAR_INPUT
      X : Real;
      X01 : Real;
      X02 : Real;
      X03 : Real;
      X04 : Real;
      X11 : Real;
      X12 : Real;
      X13 : Real;
      X14 : Real;
      X21 : Real;
      X22 : Real;
      X23 : Real;
      X24 : Real;
      X31 : Real;
      X32 : Real;
      X33 : Real;
      X34 : Real;
      L1 : Real;
      L2 : Real;
      L3 : Real;
      TC : Time;
   END_VAR
   VAR_OUTPUT
      P1 : Real;
      P2 : Real;
      P3 : Real;
      P4 : Real;
   END_VAR
   VAR
      Pset : "PARSET";
      init : Bool;
   END_VAR
BEGIN


     (* init sequence *)
     IF NOT #init THEN
       #init := TRUE;
       #Pset(TC:=#TC, X01:=#X01, X02:=#X02, X03:=#X03, X04:=#X04, X11:=#X11, X12:=#X12, X13:=#X13, X14:=#X14, X21:=#X21, X22:=#X22, X23:=#X23, X24:=#X24, X31:=#X31, X32:=#X32, X33:=#X33, X34:=#X34);
     END_IF;
     IF ABS(#X) < #L1 THEN
       #Pset(A0 := FALSE, A1 := FALSE);
     ELSIF ABS(#X) < #L2 THEN
       #Pset(A0 := TRUE, A1 := FALSE);
     ELSIF ABS(#X) < #L3 THEN
       #Pset(A0 := FALSE, A1 := TRUE);
     ELSE
       #Pset(A0 := TRUE, A1 := TRUE);
     END_IF;
     #P1 := #Pset.P1;
     #P2 := #Pset.P2;
     #P3 := #Pset.P3;
     #P4 := #Pset.P4;

   (* revision history
   hm    3.11.2007   rev 1.0
     original version

   *)
END_FUNCTION_BLOCK

FUNCTION_BLOCK "SIGNAL"   // FB215, SCL
TITLE = SIGNAL
{ S7_Optimized_Access := 'FALSE' }
AUTHOR : hugo
FAMILY : AUTOMAT
NAME : SIGNAL
VERSION : 1.0
// this function generates an output signal according to a bit pattern SIG.
// the patter is shifted to the output in time steps of TS.
// ts defaults to 128 ms if not specified.
// 
// uses: T_PLC_MS [FC64]
//       STIME [FB64],IDB_STIME [DB64]
   VAR_INPUT
      IN : Bool;
      SIG : Byte;
      TS : Time;
   END_VAR
   VAR_OUTPUT
      Q : Bool;
   END_VAR
   VAR
      tx : DWord;
      "step" : Byte;
   END_VAR
BEGIN


     IF #IN THEN
       (* an alarm is present read system time first *)
       #tx := "T_PLC_MS"();
       (* calculate the step counter which is the lowest 3 bits of (time / ts) *)
       IF #TS > t#0s THEN
         #"step" := DWORD_TO_BYTE(DINT_TO_DWORD(DWORD_TO_DINT(#tx) / T_CONV(#TS)) AND 16#0000_0007);
       ELSE
         #"step" := DWORD_TO_BYTE(SHR(IN:=#tx,N:=7) AND 16#0000_0007);
       END_IF;
       (* convert the value 0-7 in step into one bit only (bit 0-7) *)
       #"step" := SHL(IN:="one",N:=BYTE_TO_INT(#"step"));
       (* generate the output signal *)
       #Q := BYTE_TO_INT((#"step" AND #SIG)) <> 0;
     ELSE
       #Q := FALSE;
     END_IF;

   (* revision history
   hm  13.12.2007    rev 1.0
     original version

   *)
END_FUNCTION_BLOCK

FUNCTION_BLOCK "SIGNAL_4"   // FB216, SCL
TITLE = SIGNAL_4
{ S7_Optimized_Access := 'FALSE' }
AUTHOR : hugo
FAMILY : AUTOMAT
NAME : SIGNAL4
VERSION : 1.0
// this function generates one out of 4 signals specified by bit patterns S1 .. S4.
// the selected pattern will be shifted with the step time TS.
// In1 has higher priority then In2 which has higher priority then IN3 and in4 has the lowest priority.
// ts defaults to 128 ms if not specified.
// 
// uses: SIGNAL [FB215]
//       T_PLC_MS [FC64] 
//       STIME [FB64],IDB_STIME [DB64]
   VAR_INPUT
      IN1 : Bool;
      IN2 : Bool;
      IN3 : Bool;
      IN4 : Bool;
      TS : Time;
      S1 : Byte := B#16#FF;
      S2 : Byte := B#16#F0;
      S3 : Byte := B#16#AA;
      S4 : Byte := B#16#A0;
   END_VAR
   VAR_OUTPUT
      Q : Bool;
   END_VAR
   VAR
      sig : "SIGNAL";
   END_VAR
BEGIN


     (* an alarm is present read system time first *)
     (* check if an alarm is present if yes set sig to the alarm pattern otherwise exit the routine *)
     IF #IN1 THEN
       #sig(IN := TRUE, SIG := #S1, TS := #TS);
     ELSIF #IN2 THEN
       #sig(IN := TRUE, SIG := #S2, TS := #TS);
     ELSIF #IN3 THEN
       #sig(IN := TRUE, SIG := #S3, TS := #TS);
     ELSIF #IN4 THEN
       #sig(IN := TRUE, SIG := #S4, TS := #TS);
     ELSE
       #sig(IN := FALSE);
     END_IF;

     (* set the output *)
     #Q := #sig.Q;


   (* revision history
   hm  13.12.2007    rev 1.0
     original version

   *)
END_FUNCTION_BLOCK

FUNCTION_BLOCK "SRAMP"   // FB217, SCL
TITLE = SRAMP
{ S7_Optimized_Access := 'FALSE' }
AUTHOR : hugo
FAMILY : AUTOMAT
NAME : SRAMP
VERSION : 1.1
// RAMPS generates output signal which are slew rate and acceleration controlled.
// 
// uses: TC_S [FB134]
//       T_PLC_US [FC65] 
//       STIME [FB64],IDB_STIME [DB64]
   VAR_INPUT
      X : Real;
      A_UP : Real;
      A_DN : Real;
      VU_MAX : Real;
      VD_MAX : Real;
      LIMIT_HIGH : Real;
      LIMIT_LOW : Real;
      RST : Bool;
   END_VAR
   VAR_OUTPUT
      Y : Real;
      V : Real;
   END_VAR
   VAR
      cycle_time : "TC_S";
      init : Bool;
   END_VAR
BEGIN


   (* read the system_time in microseconds *)
   #cycle_time();

   (* assure range of inputs *)
   #A_UP := MAX(IN1:=0.0,IN2:=#A_UP);
   #A_DN := MIN(IN1:=0.0,IN2:=#A_DN);
   #VU_MAX := MAX(IN1:=0.0,IN2:=#VU_MAX);
   #VD_MAX := MIN(IN1:=0.0,IN2:=#VD_MAX);

   (* calculate the output offset *)
   IF #RST OR NOT #init THEN
       #init := TRUE;
       #Y := 0.0;
       #V := 0.0;
   ELSIF #X = #Y THEN
       #V := 0.0;
   ELSIF #X > #Y THEN
       (* output is too low >> ramp up and brake at the end *)
       (* accelerate the speed and limit to vu_max *)
       #V := MIN(IN1:=#V + #A_UP * #cycle_time.TC,IN2:=#VU_MAX);
       (* calculate the max speed to be able to brake and select the lowest *)
       #V := MIN(IN1:=SQRT((#Y-#X) * 2.0 * #A_DN),IN2:=#V);
       (* calculate the output and obey limits *)
       #Y := LIMIT(MN:=#LIMIT_LOW,IN:=#Y + MIN(IN1:=#V * #cycle_time.TC,IN2:=#X-#Y),MX:=#LIMIT_HIGH);
   ELSIF #X < #Y THEN
       (* output is too high >> ramp dn and brake at the end *)
       (* accelerate the speed and limit to vd_max *)
       #V := MAX(IN1:=#V + #A_DN * #cycle_time.TC,IN2:=#VD_MAX);
       (* calculate the max speed to be able to brake and select the lowest *)
       #V := MAX(IN1:=-SQRT((#Y-#X) * 2.0 * #A_UP),IN2:=#V);
       (* calculate the output and obey limits *)
       #Y := LIMIT(MN:=#LIMIT_LOW,IN:=#Y + MAX(IN1:=#V * #cycle_time.TC,IN2:=#X-#Y),MX:=#LIMIT_HIGH);
   END_IF;


   (* revision history
   hm  13. mar. 2008   rev 1.0
       original version

   hm  11. mar. 2009   rev 1.1
       real constants updated to new systax using dot

   *)
END_FUNCTION_BLOCK

FUNCTION_BLOCK "TUNE"   // FB219, SCL
TITLE = TUNE
{ S7_Optimized_Access := 'FALSE' }
AUTHOR : hugo
FAMILY : AUTOMAT
NAME : TUNE
VERSION : 1.2
// tune generates an output signal which is set by input switches.
// up to 4 switsches can be used to tune the signal up or down.
// 
// uses: T_PLC_MS [FC64]
//       STIME [FB64],IDB_STIME [DB64]
   VAR_INPUT
      SET : Bool;
      SU : Bool;
      SD : Bool;
      RST : Bool;
      SS : Real := 1.0e-1;
      Limit_L : Real;
      LIMIT_H : Real := 1.0e+2;
      RST_val : Real;
      SET_val : Real := 1.0e+2;
      T_1 : Time := T#500MS;
      T_2 : Time := T#2S;
      S1 : Real := 2.0e+0;
      S2 : Real := 1.0e+1;
   END_VAR
   VAR_OUTPUT
      Y : Real;
   END_VAR
   VAR
      tx : DWord;
      start : DWord;
      start2 : DWord;
      state : Int;
      in : Bool;
      "step" : Real;
      speed : Real;
      Y_start : Real;
      Y_start2 : Real;
   END_VAR
BEGIN


   (* read system time *)
   #tx := "T_PLC_MS"();

   IF #RST THEN
       #Y := #RST_val;
       #state := 0;
   ELSIF #SET THEN
       #Y := #SET_val;
       #state := 0;
   ELSIF #state > 0 THEN
       (* key has been pushed state machine operating *)
       (* first read the correct input *)
       IF #state = 1 THEN
           (* step up *)
           #in := #SU;
       ELSE
           (* step down *)
           #in := #SD;
       END_IF;
       (* check for single step operation *)
       IF NOT #in AND DWORD_TO_DINT(#tx) - DWORD_TO_DINT(#start) <= T_CONV(#T_1) THEN
           #Y := #Y_start + #"step";
           #state := 0;
       (* check if fast ramp needs to be generated *)
       ELSIF #in AND DWORD_TO_DINT(#tx) - DWORD_TO_DINT(#start) >= T_CONV(#T_2) THEN
           #Y := #Y_start2 + (DINT_TO_REAL(DWORD_TO_DINT(#tx) - DWORD_TO_DINT(#start2))) * #S2 / #speed;
       (* check if slow ramp needs to be generated *)
       ELSIF #in AND DWORD_TO_DINT(#tx) - DWORD_TO_DINT(#start) >= T_CONV(#T_1) THEN
           #Y := #Y_start + (DINT_TO_REAL(DWORD_TO_DINT(#tx) - DWORD_TO_DINT(#start) - T_CONV(#T_1))) * #S1 / #speed;
           #start2 := #tx;
           #Y_start2 := #Y;
       ELSIF NOT #in THEN
           #state := 0;
       END_IF;
   ELSIF #SU THEN
       (* slow step up *)
       #state := 1;
       #start := #tx;
       #"step" := #SS;
       #speed := 1000.0;
       #Y_start := #Y;
   ELSIF #SD THEN
       (* slow step down *)
       #state := 2;
       #start := #tx;
       #"step" := -#SS;
       #speed := -1000.0;
       #Y_start := #Y;
   END_IF;

   (* make sure output does not exceed limits *)
   #Y := LIMIT(MN:=#Limit_L, IN:=#Y, MX:=#LIMIT_H);


   (* revision history
   hm  3.11.2007       rev 1.0
       original version

   hm  16. mar. 2008   rev 1.1
       added type conversions to avoid warnings under codesys 3.0

   hm  11. mar. 2009   rev 1.2
       real constants updated to new systax using dot

   *)
END_FUNCTION_BLOCK

FUNCTION_BLOCK "TUNE2"   // FB220, SCL
TITLE = TUNE2
{ S7_Optimized_Access := 'FALSE' }
AUTHOR : hugo
FAMILY : AUTOMAT
NAME : TUNE2
VERSION : 1.2
// tune2 generates an output signal which is set by input switches.
// up to 4 switsches can be used to tune the signal up or down.
// 
// uses: T_PLC_MS [FC64]
//       STIME [FB64],IDB_STIME [DB64]
   VAR_INPUT
      SET : Bool;
      SU : Bool;
      SD : Bool;
      FU : Bool;
      FD : Bool;
      RST : Bool;
      SS : Real := 1.0e-1;
      FS : Real := 5.0e+0;
      Limit_L : Real;
      LIMIT_H : Real := 1.0e+2;
      RST_val : Real;
      SET_val : Real := 1.0e+2;
      TR : Time := T#500MS;
      S1 : Real := 2.0e+0;
      S2 : Real := 1.0e+1;
   END_VAR
   VAR_OUTPUT
      Y : Real;
   END_VAR
   VAR
      tx : DWord;
      start : DWord;
      state : Int;
      in : Bool;
      "step" : Real;
      speed : Real;
      Y_start : Real;
   END_VAR
BEGIN


   (* read system time *)
   #tx := "T_PLC_MS"();

   IF #RST THEN
       #Y := #RST_val;
       #state := 0;
   ELSIF #SET THEN
       #Y := #SET_val;
       #state := 0;
   ELSIF #state > 0 THEN
       (* key has been pushed state machine operating *)
       (* first read the correct input *)
       CASE #state OF
           1 : (* slow up *)
               #in := #SU;
           2 : (* slow down *)
               #in := #SD;
           3 : (* fast up *)
               #in := #FU;
           4 : (* fast down *)
               #in := #FD;
       END_CASE;
       (* check for single step operation *)
       IF NOT #in AND DWORD_TO_DINT(#tx) - DWORD_TO_DINT(#start) <= T_CONV(#TR) THEN
           #Y := #Y_start + #"step";
           #state := 0;
       (* check if ramp needs to be generated *)
       ELSIF #in AND DWORD_TO_DINT(#tx) - DWORD_TO_DINT(#start) >= T_CONV(#TR) THEN
           #Y := #Y_start + (DINT_TO_REAL(DWORD_TO_DINT(#tx) - DWORD_TO_DINT(#start) - T_CONV(#TR))) * #speed;
       ELSIF NOT #in THEN
           #state := 0;
       END_IF;
   ELSIF #SU THEN
       (* slow step up *)
       #state := 1;
       #start := #tx;
       #"step" := #SS;
       #speed := #S1 * 1.0E-3;
       #Y_start := #Y;
   ELSIF #SD THEN
       (* slow step down *)
       #state := 2;
       #start := #tx;
       #"step" := -#SS;
       #speed := -#S1 * 1.0E-3;
       #Y_start := #Y;
   ELSIF #FU THEN
       (* fast step up *)
       #state := 3;
       #start := #tx;
       #"step" := #FS;
       #speed := #S2 * 1.0E-3;
       #Y_start := #Y;
   ELSIF #FD THEN
       (* fast step down *)
       #state := 4;
       #start := #tx;
       #"step" := -#FS;
       #speed := -#S2 * 1.0E-3;
       #Y_start := #Y;
   END_IF;

   (* make sure output does not exceed limits *)
   #Y := LIMIT(MN:=#Limit_L, IN:=#Y, MX:=#LIMIT_H);


   (* revision history
   hm  3.11.2007       rev 1.0
       original version

   hm  16. 3. 2008 rev 1.1
       added type conversions to avoid warnings in codesys 3.0
       improved performance

   hm  11. mar. 2009   rev 1.2
       real constants updated to new systax using dot

   *)
END_FUNCTION_BLOCK

